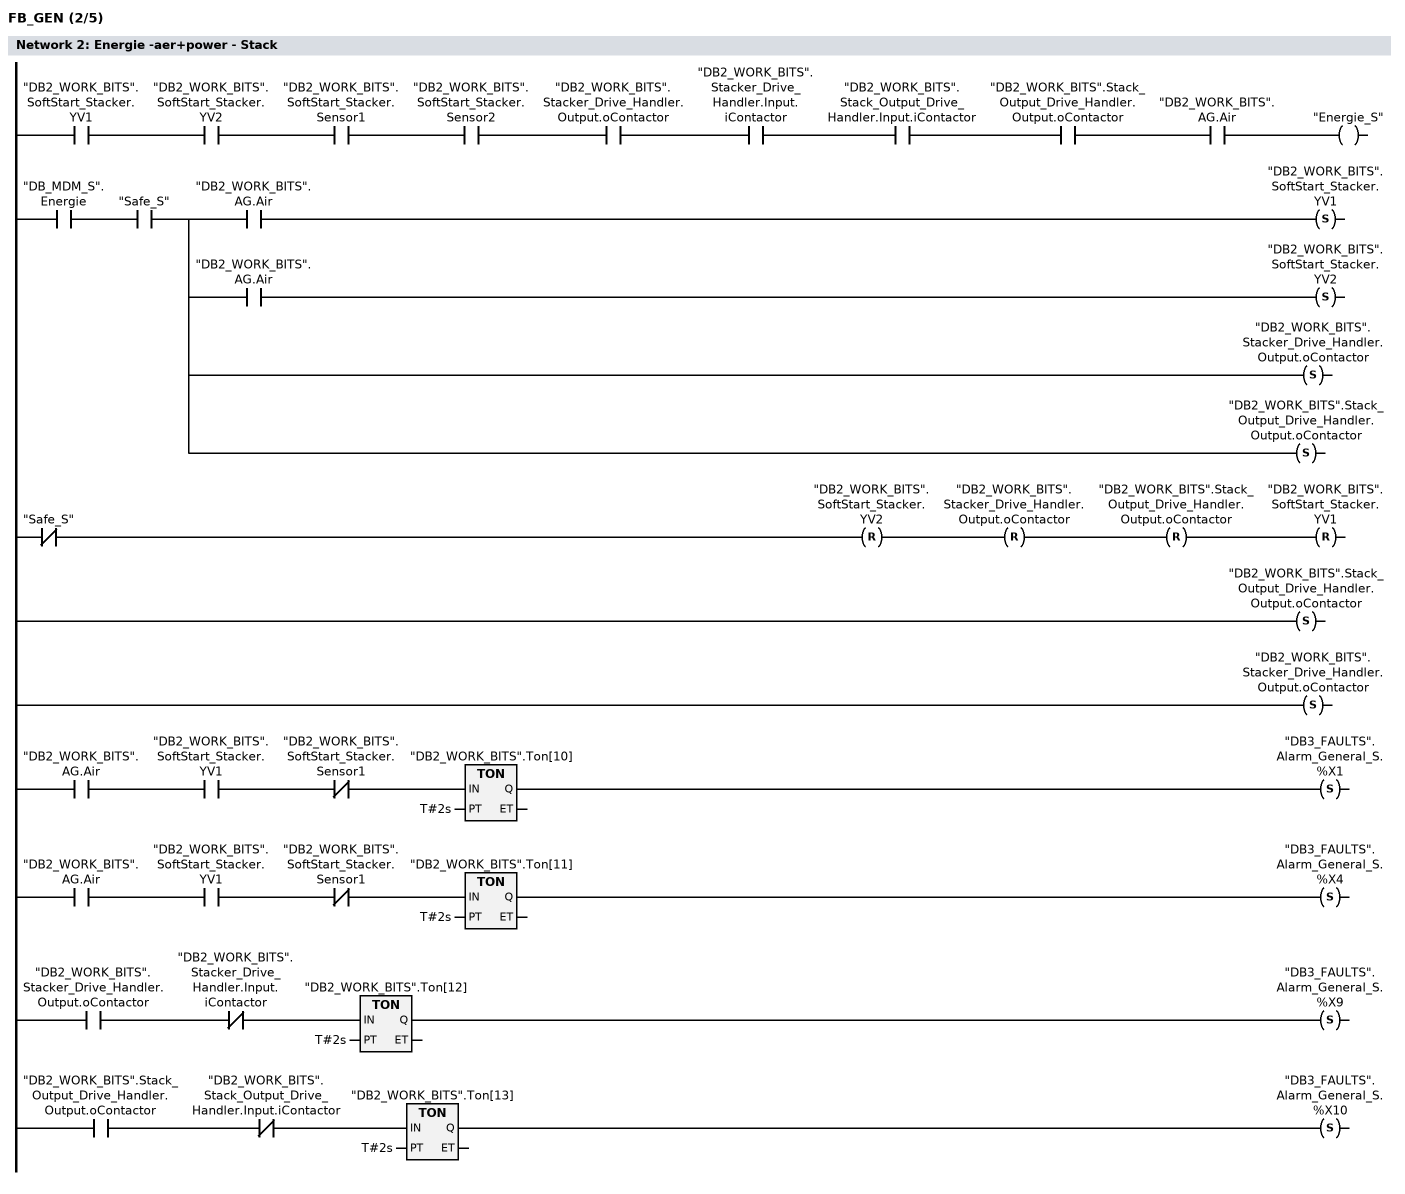
   "Energie_S" := "DB2_WORK_BITS".SoftStart_Stacker.YV1 AND "DB2_WORK_BITS".SoftStart_Stacker.YV2 AND "DB2_WORK_BITS".SoftStart_Stacker.Sensor1 AND "DB2_WORK_BITS".SoftStart_Stacker.Sensor2 AND "DB2_WORK_BITS".Stacker_Drive_Handler.Output.oContactor AND "DB2_WORK_BITS".Stacker_Drive_Handler.Input.iContactor AND "DB2_WORK_BITS".Stack_Output_Drive_Handler.Input.iContactor AND "DB2_WORK_BITS".Stack_Output_Drive_Handler.Output.oContactor AND "DB2_WORK_BITS".AG.Air;
   #_w1 := "DB_MDM_S".Energie AND "Safe_S";
   IF #_w1 AND "DB2_WORK_BITS".AG.Air THEN
       "DB2_WORK_BITS".SoftStart_Stacker.YV1 := TRUE;
       "DB2_WORK_BITS".SoftStart_Stacker.YV2 := TRUE;
   END_IF;
   IF #_w1 THEN
       "DB2_WORK_BITS".Stacker_Drive_Handler.Output.oContactor := TRUE;
       "DB2_WORK_BITS".Stack_Output_Drive_Handler.Output.oContactor := TRUE;
   END_IF;
   IF NOT "Safe_S" THEN
       "DB2_WORK_BITS".SoftStart_Stacker.YV2 := FALSE;
       "DB2_WORK_BITS".Stacker_Drive_Handler.Output.oContactor := FALSE;
       "DB2_WORK_BITS".Stack_Output_Drive_Handler.Output.oContactor := FALSE;
       "DB2_WORK_BITS".SoftStart_Stacker.YV1 := FALSE;
   END_IF;
   "DB2_WORK_BITS".Stack_Output_Drive_Handler.Output.oContactor := TRUE;
   "DB2_WORK_BITS".Stacker_Drive_Handler.Output.oContactor := TRUE;
   "DB2_WORK_BITS".Ton[10].TON(IN := "DB2_WORK_BITS".AG.Air AND "DB2_WORK_BITS".SoftStart_Stacker.YV1 AND NOT "DB2_WORK_BITS".SoftStart_Stacker.Sensor1,
                           PT := T#2s);
   IF "DB2_WORK_BITS".Ton[10].Q THEN "DB3_FAULTS".Alarm_General_S.%X1 := TRUE; END_IF;
   "DB2_WORK_BITS".Ton[11].TON(IN := "DB2_WORK_BITS".AG.Air AND "DB2_WORK_BITS".SoftStart_Stacker.YV1 AND NOT "DB2_WORK_BITS".SoftStart_Stacker.Sensor1,
                           PT := T#2s);
   IF "DB2_WORK_BITS".Ton[11].Q THEN "DB3_FAULTS".Alarm_General_S.%X4 := TRUE; END_IF;
   "DB2_WORK_BITS".Ton[12].TON(IN := "DB2_WORK_BITS".Stacker_Drive_Handler.Output.oContactor AND NOT "DB2_WORK_BITS".Stacker_Drive_Handler.Input.iContactor,
                           PT := T#2s);
   IF "DB2_WORK_BITS".Ton[12].Q THEN "DB3_FAULTS".Alarm_General_S.%X9 := TRUE; END_IF;
   "DB2_WORK_BITS".Ton[13].TON(IN := "DB2_WORK_BITS".Stack_Output_Drive_Handler.Output.oContactor AND NOT "DB2_WORK_BITS".Stack_Output_Drive_Handler.Input.iContactor,
                           PT := T#2s);
   IF "DB2_WORK_BITS".Ton[13].Q THEN "DB3_FAULTS".Alarm_General_S.%X10 := TRUE; END_IF;
END_REGION

REGION Network 3: Energie -Aer Z2_B
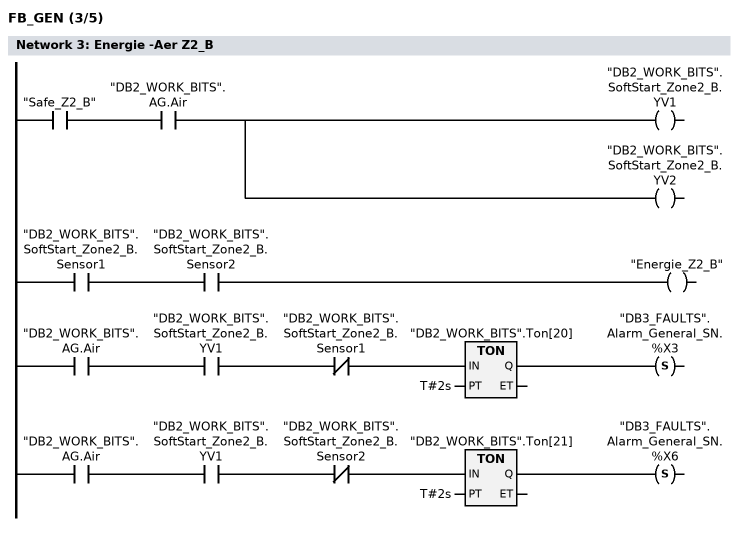
   "DB2_WORK_BITS".SoftStart_Zone2_B.YV1 := "Safe_Z2_B" AND "DB2_WORK_BITS".AG.Air;
   "DB2_WORK_BITS".SoftStart_Zone2_B.YV2 := "DB2_WORK_BITS".SoftStart_Zone2_B.YV1;
   "Energie_Z2_B" := "DB2_WORK_BITS".SoftStart_Zone2_B.Sensor1 AND "DB2_WORK_BITS".SoftStart_Zone2_B.Sensor2;
   "DB2_WORK_BITS".Ton[20].TON(IN := "DB2_WORK_BITS".AG.Air AND "DB2_WORK_BITS".SoftStart_Zone2_B.YV1 AND NOT "DB2_WORK_BITS".SoftStart_Zone2_B.Sensor1,
                           PT := T#2s);
   IF "DB2_WORK_BITS".Ton[20].Q THEN "DB3_FAULTS".Alarm_General_SN.%X3 := TRUE; END_IF;
   "DB2_WORK_BITS".Ton[21].TON(IN := "DB2_WORK_BITS".AG.Air AND "DB2_WORK_BITS".SoftStart_Zone2_B.YV1 AND NOT "DB2_WORK_BITS".SoftStart_Zone2_B.Sensor2,
                           PT := T#2s);
   IF "DB2_WORK_BITS".Ton[21].Q THEN "DB3_FAULTS".Alarm_General_SN.%X6 := TRUE; END_IF;
END_REGION

REGION Network 4: Energie -aer+power - Stack_Nou
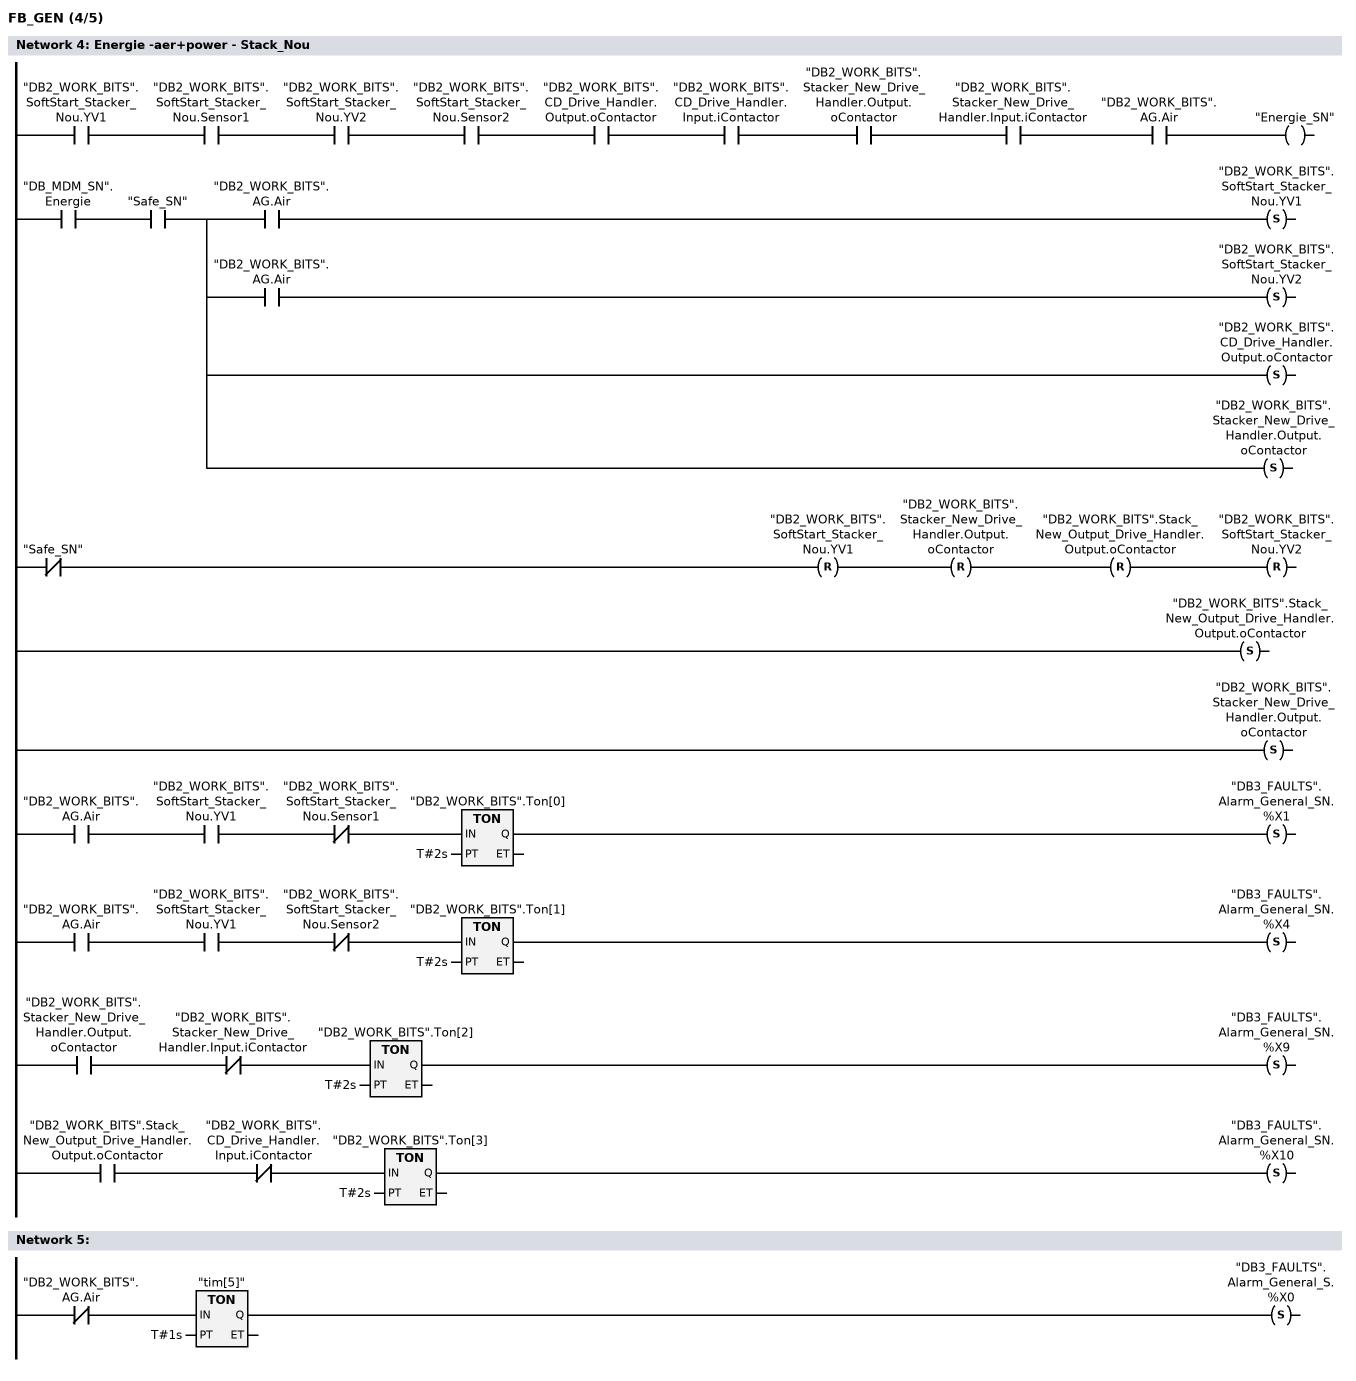
   "Energie_SN" := "DB2_WORK_BITS".SoftStart_Stacker_Nou.YV1 AND "DB2_WORK_BITS".SoftStart_Stacker_Nou.Sensor1 AND "DB2_WORK_BITS".SoftStart_Stacker_Nou.YV2 AND "DB2_WORK_BITS".SoftStart_Stacker_Nou.Sensor2 AND "DB2_WORK_BITS".CD_Drive_Handler.Output.oContactor AND "DB2_WORK_BITS".CD_Drive_Handler.Input.iContactor AND "DB2_WORK_BITS".Stacker_New_Drive_Handler.Output.oContactor AND "DB2_WORK_BITS".Stacker_New_Drive_Handler.Input.iContactor AND "DB2_WORK_BITS".AG.Air;
   #_w1 := "DB_MDM_SN".Energie AND "Safe_SN";
   IF #_w1 AND "DB2_WORK_BITS".AG.Air THEN
       "DB2_WORK_BITS".SoftStart_Stacker_Nou.YV1 := TRUE;
       "DB2_WORK_BITS".SoftStart_Stacker_Nou.YV2 := TRUE;
   END_IF;
   IF #_w1 THEN
       "DB2_WORK_BITS".CD_Drive_Handler.Output.oContactor := TRUE;
       "DB2_WORK_BITS".Stacker_New_Drive_Handler.Output.oContactor := TRUE;
   END_IF;
   IF NOT "Safe_SN" THEN
       "DB2_WORK_BITS".SoftStart_Stacker_Nou.YV1 := FALSE;
       "DB2_WORK_BITS".Stacker_New_Drive_Handler.Output.oContactor := FALSE;
       "DB2_WORK_BITS".Stack_New_Output_Drive_Handler.Output.oContactor := FALSE;
       "DB2_WORK_BITS".SoftStart_Stacker_Nou.YV2 := FALSE;
   END_IF;
   "DB2_WORK_BITS".Stack_New_Output_Drive_Handler.Output.oContactor := TRUE;
   "DB2_WORK_BITS".Stacker_New_Drive_Handler.Output.oContactor := TRUE;
   "DB2_WORK_BITS".Ton[0].TON(IN := "DB2_WORK_BITS".AG.Air AND "DB2_WORK_BITS".SoftStart_Stacker_Nou.YV1 AND NOT "DB2_WORK_BITS".SoftStart_Stacker_Nou.Sensor1,
                           PT := T#2s);
   IF "DB2_WORK_BITS".Ton[0].Q THEN "DB3_FAULTS".Alarm_General_SN.%X1 := TRUE; END_IF;
   "DB2_WORK_BITS".Ton[1].TON(IN := "DB2_WORK_BITS".AG.Air AND "DB2_WORK_BITS".SoftStart_Stacker_Nou.YV1 AND NOT "DB2_WORK_BITS".SoftStart_Stacker_Nou.Sensor2,
                           PT := T#2s);
   IF "DB2_WORK_BITS".Ton[1].Q THEN "DB3_FAULTS".Alarm_General_SN.%X4 := TRUE; END_IF;
   "DB2_WORK_BITS".Ton[2].TON(IN := "DB2_WORK_BITS".Stacker_New_Drive_Handler.Output.oContactor AND NOT "DB2_WORK_BITS".Stacker_New_Drive_Handler.Input.iContactor,
                           PT := T#2s);
   IF "DB2_WORK_BITS".Ton[2].Q THEN "DB3_FAULTS".Alarm_General_SN.%X9 := TRUE; END_IF;
   "DB2_WORK_BITS".Ton[3].TON(IN := "DB2_WORK_BITS".Stack_New_Output_Drive_Handler.Output.oContactor AND NOT "DB2_WORK_BITS".CD_Drive_Handler.Input.iContactor,
                           PT := T#2s);
   IF "DB2_WORK_BITS".Ton[3].Q THEN "DB3_FAULTS".Alarm_General_SN.%X10 := TRUE; END_IF;
END_REGION

REGION Network 5
   "tim[5]".TON(IN := NOT "DB2_WORK_BITS".AG.Air, PT := T#1s);
   IF "tim[5]".Q THEN "DB3_FAULTS".Alarm_General_S.%X0 := TRUE; END_IF;
END_REGION

REGION Network 6: rst
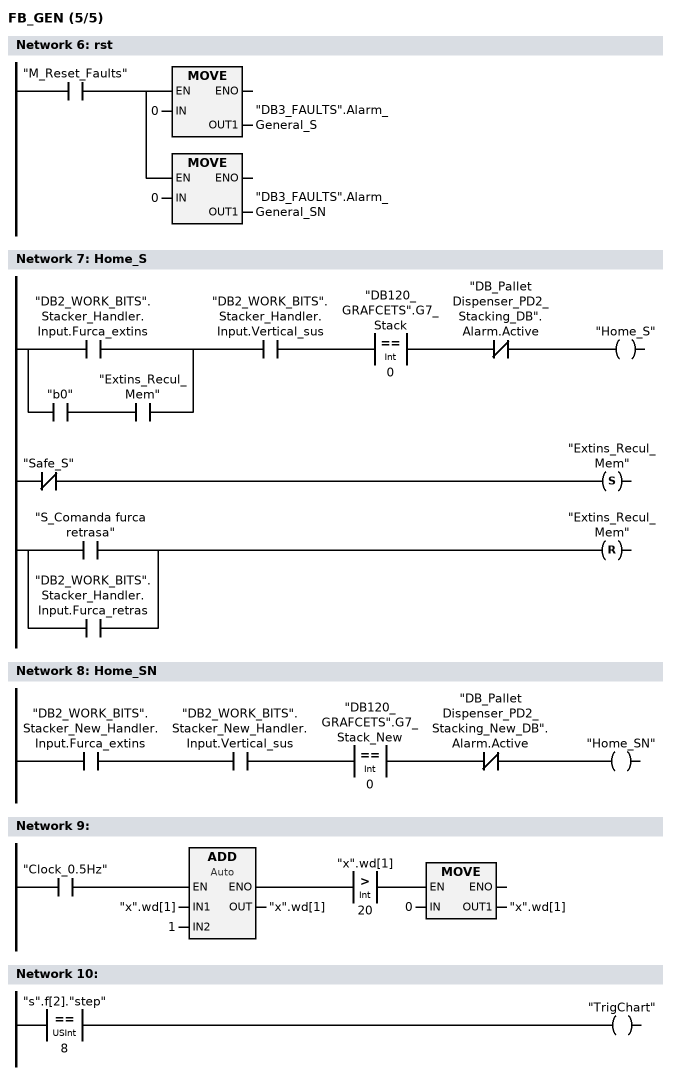
   RUNG wire#powerrail
      Contact( "M_Reset_Faults" )
      wire#w1
      Move(in := 0, out1 => "DB3_FAULTS".Alarm_General_S)
   END_RUNG
   RUNG wire#w1
      Move(in := 0, out1 => "DB3_FAULTS".Alarm_General_SN)
   END_RUNG
   // the same network as SCL:
   IF "M_Reset_Faults" THEN
       "DB3_FAULTS".Alarm_General_S := 0;
       "DB3_FAULTS".Alarm_General_SN := 0;
   END_IF;
END_REGION

REGION Network 7: Home_S
   RUNG wire#powerrail
      Contact( "DB2_WORK_BITS".Stacker_Handler.Input.Furca_extins )
      wire#w1
      Contact( "DB2_WORK_BITS".Stacker_Handler.Input.Vertical_sus )
      { S7_Templates := "SrcType := Int" } EQ_Contact(in1 := "DB120_GRAFCETS".G7_Stack, in2 := 0)
      I_Contact( "DB_PalletDispenser_PD2_Stacking_DB".Alarm.Active )
      Coil( "Home_S" )
   END_RUNG
   RUNG wire#powerrail
      Contact( "b0" )
      Contact( "Extins_Recul_Mem" )
   END_RUNG wire#w1
   RUNG wire#powerrail
      I_Contact( "Safe_S" )
      S_Coil( "Extins_Recul_Mem" )
   END_RUNG
   RUNG wire#powerrail
      Contact( "S_Comanda furca retrasa" )
      wire#w2
      R_Coil( "Extins_Recul_Mem" )
   END_RUNG
   RUNG wire#powerrail
      Contact( "DB2_WORK_BITS".Stacker_Handler.Input.Furca_retras )
   END_RUNG wire#w2
   // the same network as SCL:
   "Home_S" := ("DB2_WORK_BITS".Stacker_Handler.Input.Furca_extins OR ("b0" AND "Extins_Recul_Mem")) AND "DB2_WORK_BITS".Stacker_Handler.Input.Vertical_sus AND ("DB120_GRAFCETS".G7_Stack = 0) AND NOT "DB_PalletDispenser_PD2_Stacking_DB".Alarm.Active;
   IF NOT "Safe_S" THEN "Extins_Recul_Mem" := TRUE; END_IF;
   IF "S_Comanda furca retrasa" OR "DB2_WORK_BITS".Stacker_Handler.Input.Furca_retras THEN
       "Extins_Recul_Mem" := FALSE;
   END_IF;
END_REGION

REGION Network 8: Home_SN
   RUNG wire#powerrail
      Contact( "DB2_WORK_BITS".Stacker_New_Handler.Input.Furca_extins )
      Contact( "DB2_WORK_BITS".Stacker_New_Handler.Input.Vertical_sus )
      { S7_Templates := "SrcType := Int" } EQ_Contact(in1 := "DB120_GRAFCETS".G7_Stack_New, in2 := 0)
      I_Contact( "DB_PalletDispenser_PD2_Stacking_New_DB".Alarm.Active )
      Coil( "Home_SN" )
   END_RUNG
   // the same network as SCL:
   "Home_SN" := "DB2_WORK_BITS".Stacker_New_Handler.Input.Furca_extins AND "DB2_WORK_BITS".Stacker_New_Handler.Input.Vertical_sus AND ("DB120_GRAFCETS".G7_Stack_New = 0) AND NOT "DB_PalletDispenser_PD2_Stacking_New_DB".Alarm.Active;
END_REGION

REGION Network 9
   RUNG wire#powerrail
      Contact( "Clock_0.5Hz" )
      Add(in1 := "x".wd[1], in2 := 1, out => "x".wd[1])
      { S7_Templates := "SrcType := Int" } GT_Contact(in1 := "x".wd[1], in2 := 20)
      Move(in := 0, out1 => "x".wd[1])
   END_RUNG
   // the same network as SCL:
   IF "Clock_0.5Hz" THEN "x".wd[1] := "x".wd[1] + 1; END_IF;
   IF "Clock_0.5Hz" AND ("x".wd[1] > 20) THEN "x".wd[1] := 0; END_IF;
END_REGION

REGION Network 10
   RUNG wire#powerrail
      { S7_Templates := "SrcType := USInt" } EQ_Contact(in1 := "s".f[2]."step", in2 := 8)
      Coil( "TrigChart" )
   END_RUNG
   // the same network as SCL:
   "TrigChart" := "s".f[2]."step" = 8;
END_REGION
END_FUNCTION_BLOCK

FUNCTION_BLOCK "FB_Stack"   // FB17, LAD
{ S7_Optimized_Access := 'TRUE' }
VERSION : 0.1
   VAR_INPUT
      iEnable : Bool;
      iReset : Bool;
      iAutomatic : Bool;
      iManual : Bool;
      iManualUp : Bool;
      iManualDown : Bool;
      iManualOpenForks : Bool;
      iManualCloseForks : Bool;
      iB1_up : Bool;
      iB2_mid : Bool;
      iB10 : Bool;
      iB3_dwn : Bool;
      iB5_extins : Bool;
      iB13_retras : Bool;
      iB7_palet : Bool;
      iB8_stiva : Bool;
   END_VAR
BEGIN
END_FUNCTION_BLOCK

FUNCTION_BLOCK "FB_Init_SN"   // FB48, LAD
TITLE = td -bitii de comenzi locali (ex: #Comanda_Furca) trebuie pusi in OUT
{ S7_Optimized_Access := 'TRUE' }
VERSION : 0.1
   VAR_INPUT
      DRV : "Bits_Stacker";
   END_VAR
   VAR
      Vertical : Bool;
      Furca : Bool;
      Comanda_Furca : Bool;
      Comanda_Vertical : Bool;
      InitReq : Bool;
      Init_OK : Bool;
      Alarm_Timeout_Vertical : Bool;
      Alarm_Timeout_Furca : Bool;
      "step" : USInt;
      Init_NotPossible : Bool;
      RstStack : Bool;
      Timer_Alarms : Array[0..1] of IEC_TIMER;
   END_VAR
   VAR_TEMP   // added for the SCL form of the ladder/FBD networks
      _w1 : Bool;
      _w2 : Bool;
   END_VAR
BEGIN

REGION Network 1: ini req
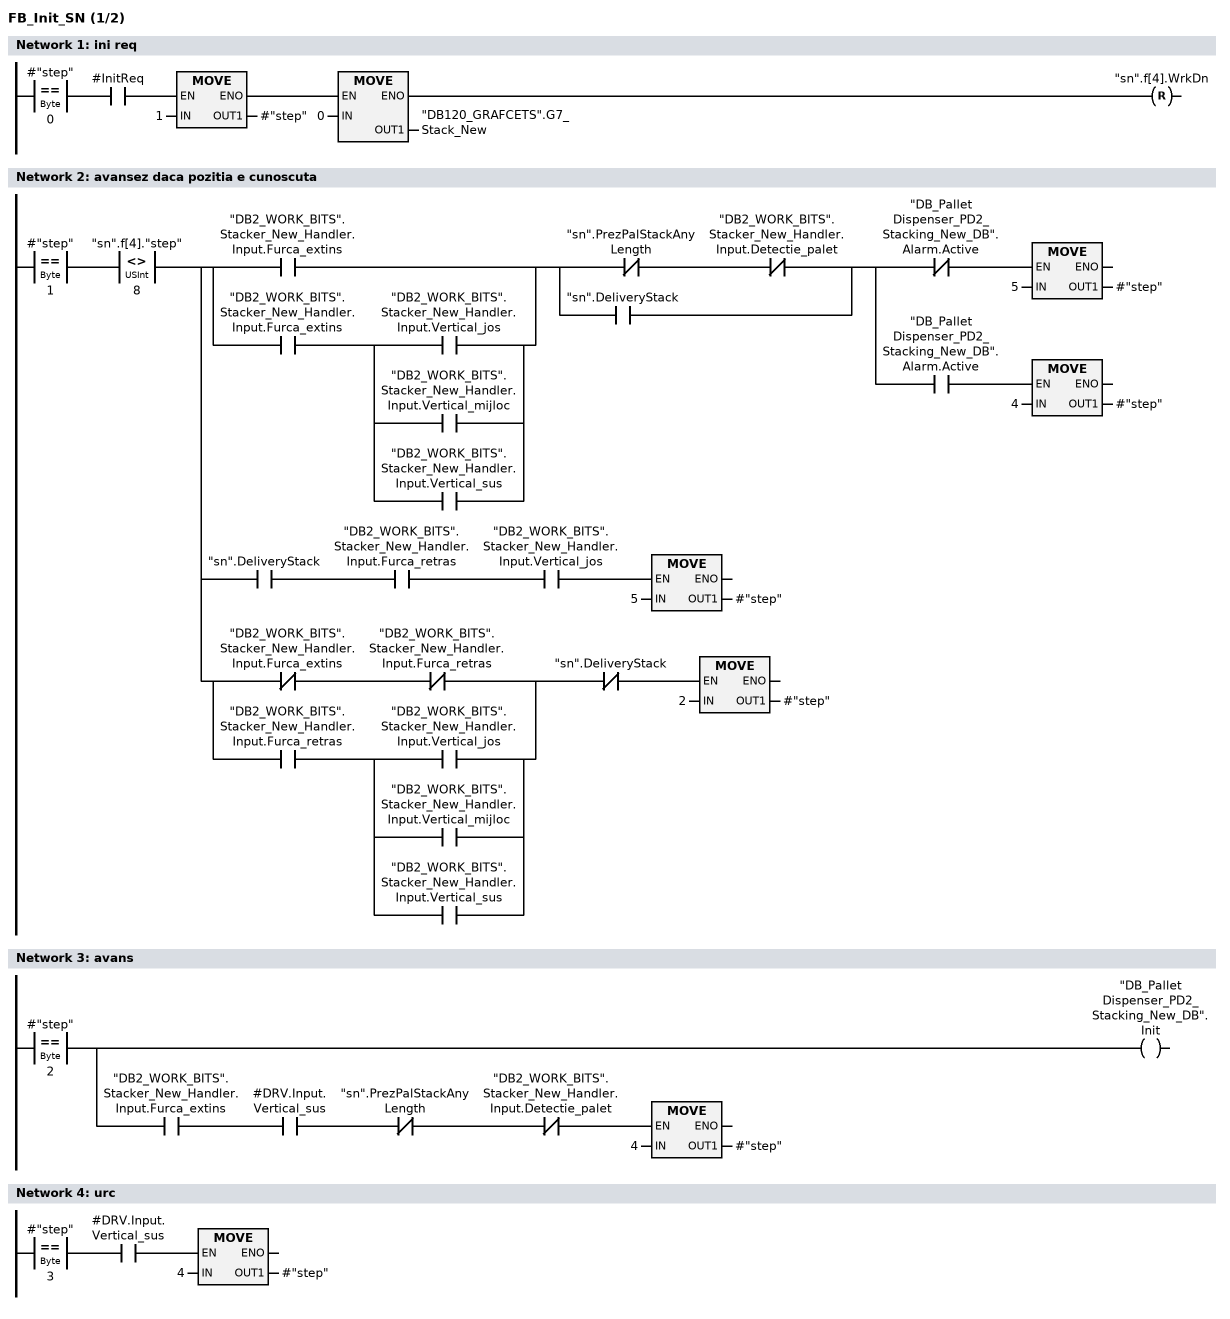
   RUNG wire#powerrail
      { S7_Templates := "SrcType := Byte" } EQ_Contact(in1 := #"step", in2 := 0)
      Contact( #InitReq )
      Move(in := 1, out1 => #"step")
      Move(in := 0, out1 => "DB120_GRAFCETS".G7_Stack_New)
      R_Coil( "sn".f[4].WrkDn )
   END_RUNG
   // the same network as SCL:
   #_w1 := (#"step" = 0) AND #InitReq;
   IF #_w1 THEN
       #"step" := 1;
       "DB120_GRAFCETS".G7_Stack_New := 0;
       "sn".f[4].WrkDn := FALSE;
   END_IF;
END_REGION

REGION Network 2: avansez daca pozitia e cunoscuta
   RUNG wire#powerrail
      { S7_Templates := "SrcType := Byte" } EQ_Contact(in1 := #"step", in2 := 1)
      { S7_Templates := "SrcType := USInt" } NE_Contact(in1 := "sn".f[4]."step", in2 := 8)
      wire#w1
      Contact( "DB2_WORK_BITS".Stacker_New_Handler.Input.Furca_extins )
      wire#w2
      I_Contact( "sn".PrezPalStackAnyLength )
      I_Contact( "DB2_WORK_BITS".Stacker_New_Handler.Input.Detectie_palet )
      wire#w4
      I_Contact( "DB_PalletDispenser_PD2_Stacking_New_DB".Alarm.Active )
      Move(in := 5, out1 => #"step")
   END_RUNG
   RUNG wire#w1
      Contact( "DB2_WORK_BITS".Stacker_New_Handler.Input.Furca_extins )
      wire#w3
      Contact( "DB2_WORK_BITS".Stacker_New_Handler.Input.Vertical_jos )
   END_RUNG wire#w2
   RUNG wire#w3
      Contact( "DB2_WORK_BITS".Stacker_New_Handler.Input.Vertical_mijloc )
   END_RUNG wire#w2
   RUNG wire#w3
      Contact( "DB2_WORK_BITS".Stacker_New_Handler.Input.Vertical_sus )
   END_RUNG wire#w2
   RUNG wire#w2
      Contact( "sn".DeliveryStack )
   END_RUNG wire#w4
   RUNG wire#w4
      Contact( "DB_PalletDispenser_PD2_Stacking_New_DB".Alarm.Active )
      Move(in := 4, out1 => #"step")
   END_RUNG
   RUNG wire#w1
      Contact( "sn".DeliveryStack )
      Contact( "DB2_WORK_BITS".Stacker_New_Handler.Input.Furca_retras )
      Contact( "DB2_WORK_BITS".Stacker_New_Handler.Input.Vertical_jos )
      Move(in := 5, out1 => #"step")
   END_RUNG
   RUNG wire#w1
      I_Contact( "DB2_WORK_BITS".Stacker_New_Handler.Input.Furca_extins )
      I_Contact( "DB2_WORK_BITS".Stacker_New_Handler.Input.Furca_retras )
      wire#w5
      I_Contact( "sn".DeliveryStack )
      Move(in := 2, out1 => #"step")
   END_RUNG
   RUNG wire#w1
      Contact( "DB2_WORK_BITS".Stacker_New_Handler.Input.Furca_retras )
      wire#w6
      Contact( "DB2_WORK_BITS".Stacker_New_Handler.Input.Vertical_jos )
   END_RUNG wire#w5
   RUNG wire#w6
      Contact( "DB2_WORK_BITS".Stacker_New_Handler.Input.Vertical_mijloc )
   END_RUNG wire#w5
   RUNG wire#w6
      Contact( "DB2_WORK_BITS".Stacker_New_Handler.Input.Vertical_sus )
   END_RUNG wire#w5
   // the same network as SCL:
   #_w1 := (#"step" = 1) AND ("sn".f[4]."step" <> 8);
   #_w2 := #_w1 AND ("DB2_WORK_BITS".Stacker_New_Handler.Input.Furca_extins OR ("DB2_WORK_BITS".Stacker_New_Handler.Input.Furca_extins AND ("DB2_WORK_BITS".Stacker_New_Handler.Input.Vertical_jos OR "DB2_WORK_BITS".Stacker_New_Handler.Input.Vertical_mijloc OR "DB2_WORK_BITS".Stacker_New_Handler.Input.Vertical_sus))) AND ((NOT "sn".PrezPalStackAnyLength AND NOT "DB2_WORK_BITS".Stacker_New_Handler.Input.Detectie_palet) OR "sn".DeliveryStack);
   IF #_w2 AND NOT "DB_PalletDispenser_PD2_Stacking_New_DB".Alarm.Active THEN #"step" := 5; END_IF;
   IF #_w2 AND "DB_PalletDispenser_PD2_Stacking_New_DB".Alarm.Active THEN #"step" := 4; END_IF;
   IF #_w1 AND "sn".DeliveryStack AND "DB2_WORK_BITS".Stacker_New_Handler.Input.Furca_retras AND "DB2_WORK_BITS".Stacker_New_Handler.Input.Vertical_jos THEN
       #"step" := 5;
   END_IF;
   IF #_w1 AND ((NOT "DB2_WORK_BITS".Stacker_New_Handler.Input.Furca_extins AND NOT "DB2_WORK_BITS".Stacker_New_Handler.Input.Furca_retras) OR ("DB2_WORK_BITS".Stacker_New_Handler.Input.Furca_retras AND ("DB2_WORK_BITS".Stacker_New_Handler.Input.Vertical_jos OR "DB2_WORK_BITS".Stacker_New_Handler.Input.Vertical_mijloc OR "DB2_WORK_BITS".Stacker_New_Handler.Input.Vertical_sus))) AND NOT "sn".DeliveryStack THEN
       #"step" := 2;
   END_IF;
END_REGION

REGION Network 3: avans
   RUNG wire#powerrail
      { S7_Templates := "SrcType := Byte" } EQ_Contact(in1 := #"step", in2 := 2)
      wire#w1
      Coil( "DB_PalletDispenser_PD2_Stacking_New_DB".Init )
   END_RUNG
   RUNG wire#w1
      Contact( "DB2_WORK_BITS".Stacker_New_Handler.Input.Furca_extins )
      Contact( #DRV.Input.Vertical_sus )
      I_Contact( "sn".PrezPalStackAnyLength )
      I_Contact( "DB2_WORK_BITS".Stacker_New_Handler.Input.Detectie_palet )
      Move(in := 4, out1 => #"step")
   END_RUNG
   // the same network as SCL:
   "DB_PalletDispenser_PD2_Stacking_New_DB".Init := #"step" = 2;
   IF "DB_PalletDispenser_PD2_Stacking_New_DB".Init AND "DB2_WORK_BITS".Stacker_New_Handler.Input.Furca_extins AND #DRV.Input.Vertical_sus AND NOT "sn".PrezPalStackAnyLength AND NOT "DB2_WORK_BITS".Stacker_New_Handler.Input.Detectie_palet THEN
       #"step" := 4;
   END_IF;
END_REGION

REGION Network 4: urc
   RUNG wire#powerrail
      { S7_Templates := "SrcType := Byte" } EQ_Contact(in1 := #"step", in2 := 3)
      Contact( #DRV.Input.Vertical_sus )
      Move(in := 4, out1 => #"step")
   END_RUNG
   // the same network as SCL:
   IF (#"step" = 3) AND #DRV.Input.Vertical_sus THEN #"step" := 4; END_IF;
END_REGION

REGION Network 5: Reset FB stacker errors
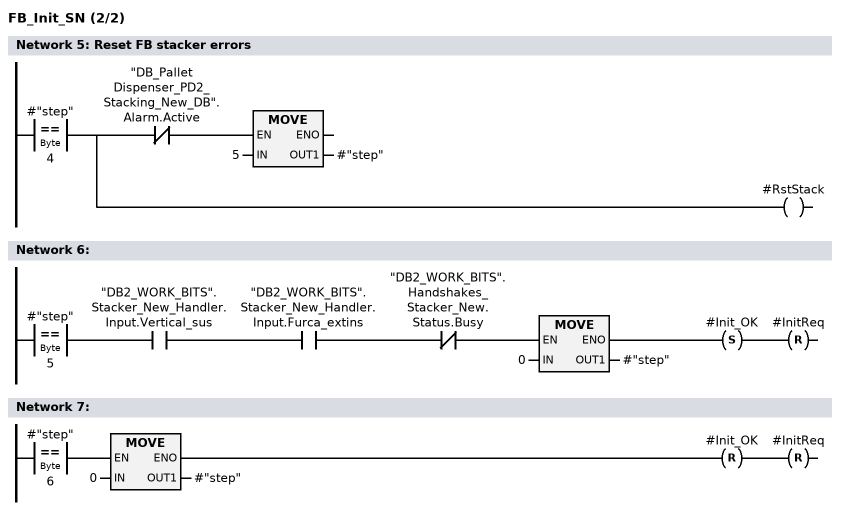
   RUNG wire#powerrail
      { S7_Templates := "SrcType := Byte" } EQ_Contact(in1 := #"step", in2 := 4)
      wire#w1
      I_Contact( "DB_PalletDispenser_PD2_Stacking_New_DB".Alarm.Active )
      Move(in := 5, out1 => #"step")
   END_RUNG
   RUNG wire#w1
      Coil( #RstStack )
   END_RUNG
   // the same network as SCL:
   #_w1 := #"step" = 4;
   IF #_w1 AND NOT "DB_PalletDispenser_PD2_Stacking_New_DB".Alarm.Active THEN #"step" := 5; END_IF;
   #RstStack := #_w1;
END_REGION

REGION Network 6
   RUNG wire#powerrail
      { S7_Templates := "SrcType := Byte" } EQ_Contact(in1 := #"step", in2 := 5)
      Contact( "DB2_WORK_BITS".Stacker_New_Handler.Input.Vertical_sus )
      Contact( "DB2_WORK_BITS".Stacker_New_Handler.Input.Furca_extins )
      I_Contact( "DB2_WORK_BITS".Handshakes_Stacker_New.Status.Busy )
      Move(in := 0, out1 => #"step")
      S_Coil( #Init_OK )
      R_Coil( #InitReq )
   END_RUNG
   // the same network as SCL:
   #_w1 := (#"step" = 5) AND "DB2_WORK_BITS".Stacker_New_Handler.Input.Vertical_sus AND "DB2_WORK_BITS".Stacker_New_Handler.Input.Furca_extins AND NOT "DB2_WORK_BITS".Handshakes_Stacker_New.Status.Busy;
   IF #_w1 THEN
       #"step" := 0;
       #Init_OK := TRUE;
       #InitReq := FALSE;
   END_IF;
END_REGION

REGION Network 7
   RUNG wire#powerrail
      { S7_Templates := "SrcType := Byte" } EQ_Contact(in1 := #"step", in2 := 6)
      Move(in := 0, out1 => #"step")
      R_Coil( #Init_OK )
      R_Coil( #InitReq )
   END_RUNG
   // the same network as SCL:
   #_w1 := #"step" = 6;
   IF #_w1 THEN
       #"step" := 0;
       #Init_OK := FALSE;
       #InitReq := FALSE;
   END_IF;
END_REGION
END_FUNCTION_BLOCK

FUNCTION_BLOCK "FB_AlarmCounter"   // FB100, SCL
{ S7_Optimized_Access := 'TRUE' }
VERSION : 0.1
   VAR_INPUT
      ResetCounters : Bool;
   END_VAR
   VAR RETAIN
      Counters : Struct
         "Destacker 110KF1 Safety Relay" : IEC_COUNTER;
         "Destacker 111KF1 Safety Barrier Relay" : IEC_COUNTER;
         "Zone 2 112KF1 Safety Relay" : IEC_COUNTER;
         "Stacker 113KF1 Safety Relay" : IEC_COUNTER;
         "Stacker 114KF1 Safety Barrier Relay 1" : IEC_COUNTER;
         "Stacker 115KF1 Safety Barrier Relay 2" : IEC_COUNTER;
         "Emergency Stop Destacker" : IEC_COUNTER;
         "Emergency Stop Zone 2" : IEC_COUNTER;
         "Emergency Stop Stacker" : IEC_COUNTER;
      END_STRUCT;
   END_VAR
BEGIN
   //count safety relay activations
   #Counters."Destacker 110KF1 Safety Relay".CTU(CU := "110KF1",
                                                 R := #ResetCounters,
                                                 PV := 0);

   #Counters."Destacker 111KF1 Safety Barrier Relay".CTU(CU := "111KF1",
                                                 R := #ResetCounters,
                                                 PV := 0);

   #Counters."Zone 2 112KF1 Safety Relay".CTU(CU := "112KF1",
                                              R := #ResetCounters,
                                              PV := 0);

   #Counters."Stacker 113KF1 Safety Relay".CTU(CU := "113KF1",
                                               R := #ResetCounters,
                                               PV := 0);

   #Counters."Stacker 114KF1 Safety Barrier Relay 1".CTU(CU := "114KF1",
                                                         R := #ResetCounters,
                                                         PV := 0);

   #Counters."Stacker 115KF1 Safety Barrier Relay 2".CTU(CU := "115KF1",
                                                         R := #ResetCounters,
                                                         PV := 0);

   #Counters."Emergency Stop Destacker".CTU(CU := "110S1",
                                            R := #ResetCounters,
                                            PV := 0);

   #Counters."Emergency Stop Zone 2".CTU(CU := "112S1",
                                         R := #ResetCounters,
                                         PV := 0);

   #Counters."Emergency Stop Stacker".CTU(CU := "113S1",
                                          R := #ResetCounters,
                                          PV := 0);
END_FUNCTION_BLOCK

FUNCTION_BLOCK "FB_IntervalTrigger"   // FB101, SCL
{ S7_Optimized_Access := 'TRUE' }
VERSION : 0.1
   VAR_OUTPUT
      bYearChanged : Bool;
      bMonthChanged : Bool;
      bWeekChanged : Bool;   // Not implemented yet
      bDayChanged : Bool;
      bHourChanged : Bool;
   END_VAR
   VAR RETAIN
      LastDay : UInt;
      LastMonth : UInt;
      LastYear : UInt;
      LastHour : UInt;
   END_VAR
   VAR
      Timer_1m : IEC_TIMER;
   END_VAR
   VAR_TEMP
      TimeDate : DTL;
      TimeDateReturn : Int;
   END_VAR
BEGIN
   #Timer_1m.TON(IN:=TRUE, PT:=T#1m);

   IF #Timer_1m.Q THEN
       #Timer_1m.IN := FALSE;
       #TimeDateReturn := RD_SYS_T(#TimeDate);
       IF #TimeDate.YEAR <> #LastYear THEN
           #bYearChanged := TRUE;
           #LastYear := #TimeDate.YEAR;
       END_IF;
       IF #TimeDate.MONTH <> #LastMonth OR #bYearChanged THEN
           #bMonthChanged := TRUE;
           #LastMonth := #TimeDate.MONTH;
       END_IF;
       IF #TimeDate.DAY <> #LastDay OR #bYearChanged  OR #bMonthChanged THEN
           #bDayChanged := TRUE;
           #LastDay := #TimeDate.DAY;
       END_IF;
       IF #TimeDate.HOUR <> #LastHour OR #bYearChanged OR #bMonthChanged OR #bDayChanged THEN
           #bHourChanged := TRUE;
           #LastHour := #TimeDate.HOUR;
       END_IF;
   ELSE
       #bHourChanged := FALSE;
       #bDayChanged := FALSE;
       #bMonthChanged := FALSE;
       #bYearChanged := FALSE;
   END_IF;
END_FUNCTION_BLOCK

FUNCTION_BLOCK "FB_EnergyCounter"   // FB102, SCL
{ S7_Optimized_Access := 'TRUE' }
VERSION : 0.1
   VAR_INPUT
      ibMeterPulse : Bool;
      ibHourChange : Bool;
      ibDayChange : Bool;
      ibMonthChange : Bool;
      ibReset : Bool;
   END_VAR
   VAR RETAIN
      Counters : Struct
         LastHour : IEC_UCOUNTER;
         LastDay : IEC_UDCOUNTER;
         LastMonth : IEC_UDCOUNTER;
      END_STRUCT;
   END_VAR
BEGIN

   #Counters.LastHour.CTU(CU := #ibMeterPulse,
                          R := #ibReset OR #ibHourChange,
                          PV := 0);

   #Counters.LastDay.CTU(CU := #ibMeterPulse,
                         R := #ibReset OR #ibDayChange,
                         PV := 0);

   #Counters.LastMonth.CTU(CU := #ibMeterPulse,
                           R := #ibReset OR #ibMonthChange,
                           PV := 0);
END_FUNCTION_BLOCK

FUNCTION_BLOCK "FB_ProductionStatistics"   // FB103, SCL
{ S7_Optimized_Access := 'TRUE' }
VERSION : 0.1
   VAR_INPUT
      ibDestroy : Bool;
      ibRepair : Bool;
      ibDayChange : Bool;
      ibMonthChange : Bool;
   END_VAR
   VAR RETAIN
      Counters : Struct
         Repairs : Struct
            LastDay : IEC_COUNTER;
            LastMonth : IEC_COUNTER;
            Repairs : Struct
               LastDay : IEC_COUNTER;
               LastMonth : IEC_COUNTER;
            END_STRUCT;
         END_STRUCT;
         Destroyed : Struct
            LastDay : IEC_COUNTER;
            LastMonth : IEC_COUNTER;
         END_STRUCT;
      END_STRUCT;
   END_VAR
   VAR
      CntPal : UInt;
      CntStack : UInt;
      CntPalS : UInt;
      fr : UInt;
      trgCntPal : Bool;
      trgCntStack : Bool;
      dat : DTL;
      dayv : UInt;
      chg_day : Bool;
   END_VAR
   VAR_TEMP
      ret : Int;
   END_VAR
BEGIN
   #Counters.Repairs.LastDay.CTU(CU := #ibRepair,
                                 R := #ibDayChange,
                                 PV := 0);

   #Counters.Repairs.LastMonth.CTU(CU := #ibRepair,
                                   R := #ibMonthChange,
                                   PV := 0);

   #Counters.Destroyed.LastDay.CTU(CU := #ibDestroy,
                                 R := #ibDayChange,
                                 PV := 0);

   #Counters.Destroyed.LastMonth.CTU(CU := #ibDestroy,
                                   R := #ibMonthChange,
                                   PV := 0);
   #ret:=RD_LOC_T(#dat);
   #chg_day := 0;
   IF #dat.DAY <> #dayv THEN
       #dayv := #dat.DAY;
       #chg_day := 1;
   END_IF;
   IF #trgCntPal THEN
       #CntPal := #CntPal + 1;
       IF #chg_day THEN
           #CntPal := 0;
       END_IF;
   END_IF;
   IF #trgCntStack THEN
       #CntStack := #CntStack + 1;
       #CntPalS := #CntPal;
       IF #chg_day THEN
           #CntStack := 0;
       END_IF;
   END_IF;
END_FUNCTION_BLOCK

FUNCTION_BLOCK "FB_PalletDispenser_PD2_Stacking"   // FB301, SCL
{ S7_Optimized_Access := 'TRUE' }